// TIA Portal project "Milk Mixing 101" (V15.1)

(* hardware
DEVICE "S7-1200 station_1"  S7-1200 Station
   slot 0: "Rack_0"  S7-1200 Rack  Rack  V1.0
   slot 1: "PLC_1"  CPU 1214C AC/DC/Rly  6ES7 214-1BG40-0XB0  V4.2
DEVICE "PC-System_1"  SIMATIC PC station
   slot 0: "SIMATIC PC station"  Rail  SIMATIC PC-Station  V1.0
      slot 125: "Stationmanager"  Station_Manager  V6.0.4
   slot 1: "HMI_RT_1"  WinCC RT Advanced  6AV2 104-0xxxx-xxxx  15.1.0.0
      slot 33792: "Host interface"  Host interface
   slot 2: "IE general_1"  IE General  IE_CP  V8.2.0
*)

// ===== PLC "PLC_1"  CPU 1214C AC/DC/Rly =====

VAR_GLOBAL   // PLC tag table "Default tag table"
   "Auto_Start" AT %M0.0 : Bool;
   "Param_set" AT %M0.1 : Bool;
   "Timer_T123_ET" AT %MD0 : Time;
   "Filling_T123_Done" AT %M4.0 : Bool;
   "Filling_W1_Done" AT %M4.1 : Bool;
   "Mixing_Done" AT %M4.2 : Bool;
   "Pumping_Done" AT %M4.3 : Bool;
   "Pastorizing_Done" AT %M4.4 : Bool;
   "Filler_Done" AT %M4.5 : Bool;
   "MoveFork" AT %MD4 : DWord;
END_VAR

DATA_BLOCK "Recipe_Params"   // DB1
{ S7_Optimized_Access := 'TRUE' }
VERSION : 0.1
   VAR
      Flavour_Vol : Real;
      Milk_Vol : Real;
      Mixing_time : Time;
      Pastorizing_time : Time;
      Pastorizing_temp : Real;
      Filling_speed : Real;
      Flavour : Int;
   END_VAR
BEGIN
END_DATA_BLOCK

DATA_BLOCK "Devices"   // DB2
{ S7_Optimized_Access := 'TRUE' }
VERSION : 0.1
   VAR
      V11 : Bool;
      V12 : Bool;
      V13 : Bool;
      T1 : Bool;
      T2 : Bool;
      T3 : Bool;
      V21 : Bool;
      V22 : Bool;
      V23 : Bool;
      Mixer : Bool;
      W1 : Bool;
      V3 : Bool;
      Pump : Bool;
      V4 : Bool;
      Pastrorizer : Bool;
      v5 : Bool;
      Filler : Bool;
      Fork_Lift : Bool;
   END_VAR
BEGIN
END_DATA_BLOCK

DATA_BLOCK "SCADA_inputs"   // DB3
{ S7_Optimized_Access := 'TRUE' }
VERSION : 0.1
   VAR
      Start : Bool;
      Stop : Bool;
      Auto_On : Bool;
   END_VAR
BEGIN
END_DATA_BLOCK

DATA_BLOCK "Timer_ET"   // DB5
{ S7_Optimized_Access := 'TRUE' }
VERSION : 0.1
   VAR
      FillingTanks_ET : Time;
      FillingW1_ET : Time;
      MixingTimer_ET : Time;
      PumpingTimer_ET : Time;
      pastorizingTimer_ET : Time;
      FillerTimer_ET : Time;
   END_VAR
BEGIN
END_DATA_BLOCK

// folder: System blocks/Program resources

DATA_BLOCK "Filling_T1_2_3"   // DB4
{ S7_Optimized_Access := 'TRUE' }
AUTHOR : Simatic
FAMILY : IEC
NAME : IEC_TMR
VERSION : 1.0
// stored: InstanceOfName IEC_TIMER
"IEC_TIMER"
BEGIN
END_DATA_BLOCK

DATA_BLOCK "Filling_W1"   // DB6
{ S7_Optimized_Access := 'TRUE' }
AUTHOR : Simatic
FAMILY : IEC
NAME : IEC_TMR
VERSION : 1.0
// stored: InstanceOfName IEC_TIMER
"IEC_TIMER"
BEGIN
END_DATA_BLOCK

DATA_BLOCK "Mixing_timer"   // DB7
{ S7_Optimized_Access := 'TRUE' }
AUTHOR : Simatic
FAMILY : IEC
NAME : IEC_TMR
VERSION : 1.0
// stored: InstanceOfName IEC_TIMER
"IEC_TIMER"
BEGIN
END_DATA_BLOCK

DATA_BLOCK "Pumping_Timer"   // DB8
{ S7_Optimized_Access := 'TRUE' }
AUTHOR : Simatic
FAMILY : IEC
NAME : IEC_TMR
VERSION : 1.0
// stored: InstanceOfName IEC_TIMER
"IEC_TIMER"
BEGIN
END_DATA_BLOCK

DATA_BLOCK "Pastorizing_timer"   // DB9
{ S7_Optimized_Access := 'TRUE' }
AUTHOR : Simatic
FAMILY : IEC
NAME : IEC_TMR
VERSION : 1.0
// stored: InstanceOfName IEC_TIMER
"IEC_TIMER"
BEGIN
END_DATA_BLOCK

DATA_BLOCK "Filler_Timer"   // DB10
{ S7_Optimized_Access := 'TRUE' }
AUTHOR : Simatic
FAMILY : IEC
NAME : IEC_TMR
VERSION : 1.0
// stored: InstanceOfName IEC_TIMER
"IEC_TIMER"
BEGIN
END_DATA_BLOCK

DATA_BLOCK "Move_Fork"   // DB11
{ S7_Optimized_Access := 'TRUE' }
AUTHOR : Simatic
FAMILY : IEC
NAME : IEC_TMR
VERSION : 1.0
// stored: InstanceOfName IEC_TIMER
"IEC_TIMER"
BEGIN
END_DATA_BLOCK

// folder: (top level)

ORGANIZATION_BLOCK "Main"   // OB1, LAD, ProgramCycle
TITLE = "Main Program Sweep (Cycle)"
{ S7_Optimized_Access := 'TRUE' }
VERSION : 0.1
   VAR_INPUT
      Initial_Call : Bool;   // Initial call of this OB
      Remanence : Bool;   // =True, if remanent data are available
   END_VAR
BEGIN

REGION Network 1: Starting in Auto Mode
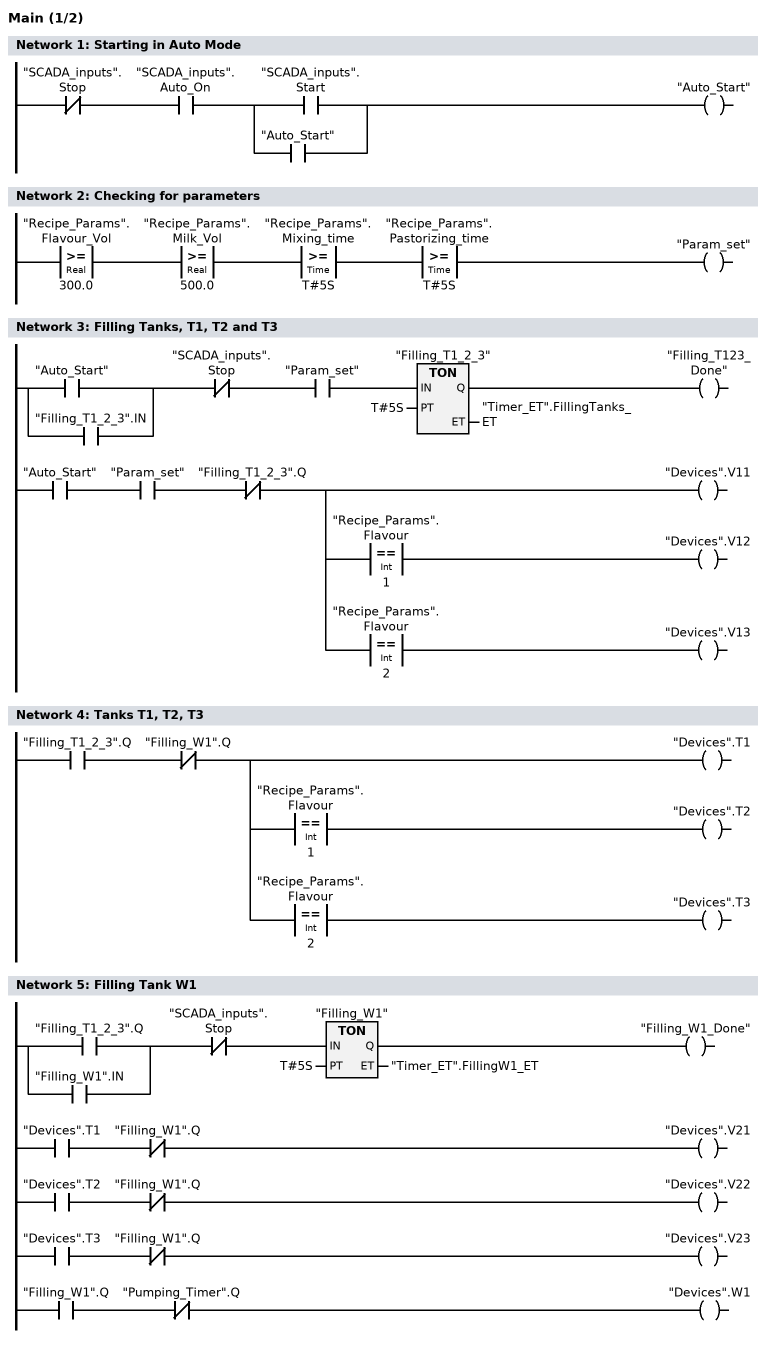
   RUNG wire#powerrail
      I_Contact( "SCADA_inputs".Stop )
      Contact( "SCADA_inputs".Auto_On )
      wire#w1
      Contact( "SCADA_inputs".Start )
      wire#w2
      Coil( "Auto_Start" )
   END_RUNG
   RUNG wire#w1
      Contact( "Auto_Start" )
   END_RUNG wire#w2
   // the same network as SCL:
   "Auto_Start" := NOT "SCADA_inputs".Stop AND "SCADA_inputs".Auto_On AND ("SCADA_inputs".Start OR "Auto_Start");
END_REGION

REGION Network 2: Checking for parameters
   RUNG wire#powerrail
      { S7_Templates := "SrcType := Real" } GE_Contact(in1 := "Recipe_Params".Flavour_Vol, in2 := 300.0)
      { S7_Templates := "SrcType := Real" } GE_Contact(in1 := "Recipe_Params".Milk_Vol, in2 := 500.0)
      { S7_Templates := "SrcType := Time" } GE_Contact(in1 := "Recipe_Params".Mixing_time, in2 := T#5S)
      { S7_Templates := "SrcType := Time" } GE_Contact(in1 := "Recipe_Params".Pastorizing_time, in2 := T#5S)
      Coil( "Param_set" )
   END_RUNG
   // the same network as SCL:
   "Param_set" := ("Recipe_Params".Flavour_Vol >= 300.0) AND ("Recipe_Params".Milk_Vol >= 500.0) AND ("Recipe_Params".Mixing_time >= T#5S) AND ("Recipe_Params".Pastorizing_time >= T#5S);
END_REGION

REGION Network 3: Filling Tanks, T1, T2 and T3
   "Filling_T1_2_3".TON(IN := ("Auto_Start" OR "Filling_T1_2_3".IN) AND NOT "SCADA_inputs".Stop AND "Param_set",
                        PT := T#5S,
                        ET => "Timer_ET".FillingTanks_ET);
   "Filling_T123_Done" := "Filling_T1_2_3".Q;
   "Devices".V11 := "Auto_Start" AND "Param_set" AND NOT "Filling_T1_2_3".Q;
   "Devices".V12 := "Devices".V11 AND ("Recipe_Params".Flavour = 1);
   "Devices".V13 := "Devices".V11 AND ("Recipe_Params".Flavour = 2);
END_REGION

REGION Network 4: Tanks T1, T2, T3
   RUNG wire#powerrail
      Contact( "Filling_T1_2_3".Q )
      I_Contact( "Filling_W1".Q )
      wire#w1
      Coil( "Devices".T1 )
   END_RUNG
   RUNG wire#w1
      { S7_Templates := "SrcType := Int" } EQ_Contact(in1 := "Recipe_Params".Flavour, in2 := 1)
      Coil( "Devices".T2 )
   END_RUNG
   RUNG wire#w1
      { S7_Templates := "SrcType := Int" } EQ_Contact(in1 := "Recipe_Params".Flavour, in2 := 2)
      Coil( "Devices".T3 )
   END_RUNG
   // the same network as SCL:
   "Devices".T1 := "Filling_T1_2_3".Q AND NOT "Filling_W1".Q;
   "Devices".T2 := "Devices".T1 AND ("Recipe_Params".Flavour = 1);
   "Devices".T3 := "Devices".T1 AND ("Recipe_Params".Flavour = 2);
END_REGION

REGION Network 5: Filling Tank W1
   "Filling_W1".TON(IN := ("Filling_T1_2_3".Q OR "Filling_W1".IN) AND NOT "SCADA_inputs".Stop,
                    PT := T#5S,
                    ET => "Timer_ET".FillingW1_ET);
   "Filling_W1_Done" := "Filling_W1".Q;
   "Devices".V21 := "Devices".T1 AND NOT "Filling_W1".Q;
   "Devices".V22 := "Devices".T2 AND NOT "Filling_W1".Q;
   "Devices".V23 := "Devices".T3 AND NOT "Filling_W1".Q;
   "Devices".W1 := "Filling_W1".Q AND NOT "Pumping_Timer".Q;
END_REGION

REGION Network 6: Mixing
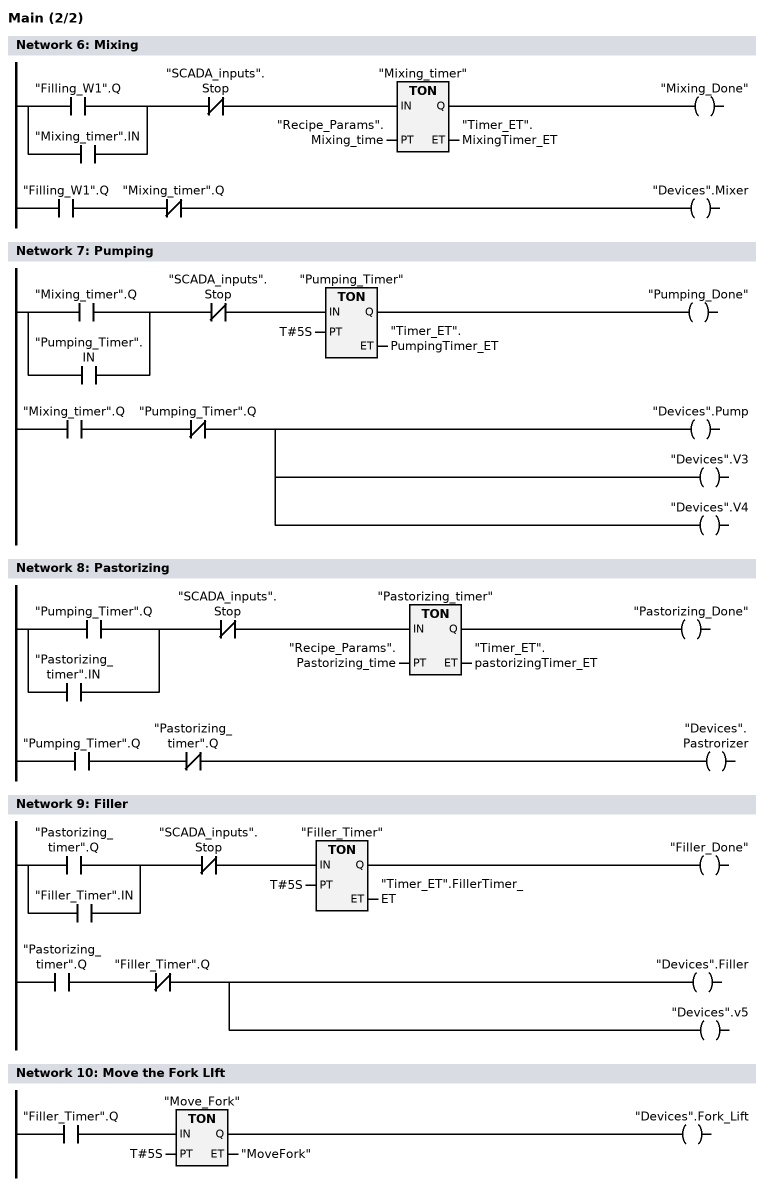
   "Mixing_timer".TON(IN := ("Filling_W1".Q OR "Mixing_timer".IN) AND NOT "SCADA_inputs".Stop,
                      PT := "Recipe_Params".Mixing_time,
                      ET => "Timer_ET".MixingTimer_ET);
   "Mixing_Done" := "Mixing_timer".Q;
   "Devices".Mixer := "Filling_W1".Q AND NOT "Mixing_timer".Q;
END_REGION

REGION Network 7: Pumping
   "Pumping_Timer".TON(IN := ("Mixing_timer".Q OR "Pumping_Timer".IN) AND NOT "SCADA_inputs".Stop,
                       PT := T#5S,
                       ET => "Timer_ET".PumpingTimer_ET);
   "Pumping_Done" := "Pumping_Timer".Q;
   "Devices".Pump := "Mixing_timer".Q AND NOT "Pumping_Timer".Q;
   "Devices".V3 := "Devices".Pump;
   "Devices".V4 := "Devices".Pump;
END_REGION

REGION Network 8: Pastorizing
   "Pastorizing_timer".TON(IN := ("Pumping_Timer".Q OR "Pastorizing_timer".IN) AND NOT "SCADA_inputs".Stop,
                           PT := "Recipe_Params".Pastorizing_time,
                           ET => "Timer_ET".pastorizingTimer_ET);
   "Pastorizing_Done" := "Pastorizing_timer".Q;
   "Devices".Pastrorizer := "Pumping_Timer".Q AND NOT "Pastorizing_timer".Q;
END_REGION

REGION Network 9: Filler
   "Filler_Timer".TON(IN := ("Pastorizing_timer".Q OR "Filler_Timer".IN) AND NOT "SCADA_inputs".Stop,
                      PT := T#5S,
                      ET => "Timer_ET".FillerTimer_ET);
   "Filler_Done" := "Filler_Timer".Q;
   "Devices".Filler := "Pastorizing_timer".Q AND NOT "Filler_Timer".Q;
   "Devices".v5 := "Devices".Filler;
END_REGION

REGION Network 10: Move the Fork LIft
   "Move_Fork".TON(IN := "Filler_Timer".Q, PT := T#5S, ET => "MoveFork");
   "Devices".Fork_Lift := "Move_Fork".Q;
END_REGION
END_ORGANIZATION_BLOCK

(* ===== HMI "HMI_RT_1" =====
system functions are stored by id; their names below are inferred from use
connection "HMI_Connection_1": ETHERNET, S7_1200_OMS

HMI tags "Default tag table"
   "Recipe_Params_Flavour" : Int = PLC Recipe_Params.Flavour, 1 s
   "Recipe_Params_Flavour_Vol" : Real = PLC Recipe_Params.Flavour_Vol, 1 s
   "Recipe_Params_Milk_Vol" : Real = PLC Recipe_Params.Milk_Vol, 1 s
   "Recipe_Params_Mixing_time" : Time = PLC Recipe_Params.Mixing_time, 1 s
   "Recipe_Params_Pastorizing_time" : Time = PLC Recipe_Params.Pastorizing_time, 1 s
   "Recipe_Params_Pastorizing_temp" : Real = PLC Recipe_Params.Pastorizing_temp, 1 s
   "Recipe_Params_Filling_speed" : Real = PLC Recipe_Params.Filling_speed, 1 s
   "SCADA_inputs_Start" : Bool = PLC SCADA_inputs.Start, 1 s
   "SCADA_inputs_Stop" : Bool = PLC SCADA_inputs.Stop, 1 s
   "SCADA_inputs_Auto_On" : Bool = PLC SCADA_inputs.Auto_On, 1 s
   "Devices_V11" : Bool = PLC Devices.V11, 1 s
   "Devices_V12" : Bool = PLC Devices.V12, 1 s
   "Devices_V13" : Bool = PLC Devices.V13, 1 s
   "Devices_T1" : Bool = PLC Devices.T1, 1 s
   "Devices_T2" : Bool = PLC Devices.T2, 1 s
   "Devices_T3" : Bool = PLC Devices.T3, 1 s
   "Devices_V21" : Bool = PLC Devices.V21, 1 s
   "Devices_V22" : Bool = PLC Devices.V22, 1 s
   "Devices_V23" : Bool = PLC Devices.V23, 1 s
   "Devices_Mixer" : Bool = PLC Devices.Mixer, 1 s
   "Devices_W1" : Bool = PLC Devices.W1, 1 s
   "Devices_V3" : Bool = PLC Devices.V3, 1 s
   "Devices_Pump" : Bool = PLC Devices.Pump, 1 s
   "Devices_V4" : Bool = PLC Devices.V4, 1 s
   "Devices_Pastrorizer" : Bool = PLC Devices.Pastrorizer, 1 s
   "Devices_v5" : Bool = PLC Devices.v5, 1 s
   "Devices_Filler" : Bool = PLC Devices.Filler, 1 s
   "MoveFork" : DWord = PLC MoveFork AT %MD4, 1 s
   "Timer_ET_FillingW1_ET" : Time = PLC Timer_ET.FillingW1_ET, 1 s
   "Auto_Start" : Bool = PLC Auto_Start AT %M0.0, 1 s

text list "Flavour": 1 'Strawberry'; 2 'Chocolate'

screen "Main_Screen" 1920x1068
   TextField "Text field_1" at 647,26 size 456x34; Text 'MILK MIXING SYSTEM'
   SymbolLibrary "Symbol library_1" at 52,135 size 108x126
   SymbolLibrary "Symbol library_2" at 254,136 size 108x126
   SymbolLibrary "Symbol library_3" at 459,136 size 108x126
   SymbolLibrary "Symbol library_4" at 66,359 size 85x71
      Appearance <- "Devices_T1"
   SymbolLibrary "Symbol library_5" at 267,356 size 85x71
      Appearance <- "Devices_T2"
   SymbolLibrary "Symbol library_6" at 471,360 size 85x71
      Appearance <- "Devices_T3"
   SymbolLibrary "Symbol library_7" at 98,262 size 16x99
      Appearance <- "Devices_V11"
   SymbolLibrary "Symbol library_8" at 300,262 size 16x99
      Appearance <- "Devices_V12"
   SymbolLibrary "Symbol library_9" at 507,261 size 16x99
      Appearance <- "Devices_V13"
   SymbolLibrary "Symbol library_10" at 77,292 size 38x41
      Appearance <- "Devices_V11"
   SymbolLibrary "Symbol library_11" at 280,290 size 38x41
      Appearance <- "Devices_V12"
   SymbolLibrary "Symbol library_12" at 487,292 size 38x41
      Appearance <- "Devices_V13"
   SymbolLibrary "Symbol library_13" at 211,552 size 201x153
      Appearance <- "Devices_W1"
   SymbolLibrary "Symbol library_14" at 100,425 size 16x84
      Appearance <- "Devices_V21"
   SymbolLibrary "Symbol library_15" at 302,426 size 16x130
      Appearance <- "Devices_V22"
   SymbolLibrary "Symbol library_16" at 506,430 size 16x76
      Appearance <- "Devices_V23"
   SymbolLibrary "Symbol library_17" at 384,517 size 103x16
      Appearance <- "Devices_V23"
   SymbolLibrary "Symbol library_18" at 133,518 size 83x16
      Appearance <- "Devices_V21"
   SymbolLibrary "Symbol library_19" at 352,516 size 33x35
   SymbolLibrary "Symbol library_20" at 213,517 size 29x38
   SymbolLibrary "Symbol library_21" at 99,505 size 35x27
   SymbolLibrary "Symbol library_22" at 486,502 size 36x30
   SymbolLibrary "Symbol library_23" at 525,809 size 101x89
      Appearance <- "Devices_Pump"
   SymbolLibrary "Symbol library_25" at 299,704 size 23x120
      Appearance <- "Devices_V3"
   SymbolLibrary "Symbol library_26" at 339,842 size 188x17
      Appearance <- "Devices_V3"
   SymbolLibrary "Symbol library_24" at 416,812 size 43x49
      Appearance <- "Devices_V3"
   SymbolLibrary "Symbol library_27" at 299,823 size 42x37
   SymbolLibrary "Symbol library_28" at 822,414 size 120x120
      Appearance <- "Devices_Pastrorizer"
   SymbolLibrary "Symbol library_29" at 713,502 size 18x301
      Appearance <- "Devices_V4"
   SymbolLibrary "Symbol library_30" at 626,818 size 59x20
   SymbolLibrary "Symbol library_31" at 751,466 size 76x19
      Appearance <- "Devices_V4"
   SymbolLibrary "Symbol library_32" at 712,466 size 39x39
   SymbolLibrary "Symbol library_33" at 685,801 size 49x36
   SymbolLibrary "Symbol library_34" at 762,436 size 43x49
      Appearance <- "Devices_V4"
   SymbolLibrary "Symbol library_35" at 858,678 size 120x120
      Appearance <- "Devices_Filler"
   SymbolLibrary "Symbol library_36" at 869,522 size 21x157
      Appearance <- "Devices_v5"
   SymbolLibrary "Symbol library_37" at 832,582 size 64x35
      Appearance <- "Devices_v5"
   SymbolLibrary "Symbol library_38" at 973,755 size 239x43
   SymbolLibrary "Symbol library_39" at 1206,691 size 120x120
      HorizontalMovement <- "MoveFork"
   Switch "Switch_1" at 1130,109 size 108x55; CaptionText 'MODE'; TextOff 'MANUAL'; TextOn 'AUTO'
      on SwitchOn: SetBit("SCADA_inputs_Auto_On")
      on SwitchOff: ResetBit("SCADA_inputs_Auto_On")
   Button "Button_1" at 1285,129 size 96x32; TextOff 'START'
      on Press: SetBit("SCADA_inputs_Start")
      on Release: ResetBit("SCADA_inputs_Start")
   Button "Button_2" at 1437,130 size 96x32; TextOff 'STOP'
      on Press: SetBit("SCADA_inputs_Stop")
      on Release: ResetBit("SCADA_inputs_Stop")
   TextField "Text field_2" at 1221,197 size 321x27; Text 'Recipe Parameter'
   TextField "Text field_3" at 1149,278 size 115x22; Text 'Flavour'
   TextField "Text field_4" at 1137,338 size 179x22; Text 'Flavour Volume'
   TextField "Text field_5" at 1140,386 size 159x22; Text 'Milk Volume'
   TextField "Text field_6" at 1138,426 size 155x22; Text 'Mixing Time'
   TextField "Text field_7" at 1134,470 size 185x22; Text 'Pastorizing Time'
   TextField "Text field_8" at 1135,515 size 198x22; Text 'Pastorizing Temp'
   TextField "Text field_9" at 1141,560 size 182x22; Text 'Filling Speed'
   SymbolicIOField "Symbolic I/O field_1" at 1294,277 size 142x33; TextOff '0'; TextOn '1'; TextList "Flavour"
      ProcessValue <- "Recipe_Params_Flavour"
      Visibility <- "Auto_Start"
   IOField "I/O field_1" at 1296,333 size 96x32; FormatPattern 9999
      ProcessValue <- "Recipe_Params_Flavour_Vol"
      Visibility <- "Auto_Start"
   IOField "I/O field_2" at 1296,382 size 96x32; FormatPattern 9999
      ProcessValue <- "Recipe_Params_Milk_Vol"
      Visibility <- "Auto_Start"
   IOField "I/O field_3" at 1296,422 size 96x32; FormatPattern 99999
      ProcessValue <- "Recipe_Params_Mixing_time"
      Visibility <- "Auto_Start"
   IOField "I/O field_4" at 1297,466 size 96x32; FormatPattern 99999
      ProcessValue <- "Recipe_Params_Pastorizing_time"
      Visibility <- "Auto_Start"
   IOField "I/O field_5" at 1298,511 size 96x32; FormatPattern 9999
      ProcessValue <- "Recipe_Params_Pastorizing_temp"
      Visibility <- "Auto_Start"
   IOField "I/O field_6" at 1297,558 size 96x32; FormatPattern 9999
      ProcessValue <- "Recipe_Params_Filling_speed"
      Visibility <- "Auto_Start"
   TextField "Text field_10" at 1415,337 size 53x22; Text 'ltr'
   TextField "Text field_11" at 1412,382 size 56x22; Text 'ltr'
   TextField "Text field_12" at 1410,426 size 77x22; Text 'ms'
   TextField "Text field_13" at 1408,476 size 87x22; Text 'ms'
   TextField "Text field_14" at 1413,516 size 81x22; Text 'c'
   TextField "Text field_15" at 1399,560 size 177x22; Text 'Bottle/min'
   TextField "Text field_16" at 43,300 size 35x22; Text 'V11'
   TextField "Text field_17" at 245,300 size 35x22; Text 'V12'
   TextField "Text field_18" at 453,302 size 35x22; Text 'V13'
   TextField "Text field_19" at 100,376 size 24x22; Text 'T1'
   TextField "Text field_20" at 302,372 size 24x22; Text 'T2'
   TextField "Text field_21" at 498,376 size 24x22; Text 'T3'
   SymbolLibrary "Symbol library_40" at 73,454 size 47x35
      Appearance <- "Devices_V21"
   SymbolLibrary "Symbol library_41" at 272,457 size 47x35
      Appearance <- "Devices_V22"
   SymbolLibrary "Symbol library_42" at 478,457 size 47x35
      Appearance <- "Devices_V23"
   TextField "Text field_22" at 40,461 size 35x22; Text 'V21'
   TextField "Text field_23" at 237,464 size 35x22; Text 'V22'
   TextField "Text field_24" at 443,467 size 35x22; Text 'V23'
   TextField "Text field_25" at 289,657 size 30x22; Text 'W1'
   SymbolLibrary "Symbol library_43" at 240,519 size 73x75
      Appearance <- "Devices_Mixer"
   TextField "Text field_26" at 257,600 size 48x22; Text 'Mixer'
   TextField "Text field_27" at 423,790 size 25x22; Text 'V3'
   TextField "Text field_28" at 770,415 size 25x22; Text 'V4'
   TextField "Text field_29" at 546,787 size 46x22; Text 'Pump'
   TextField "Text field_30" at 827,393 size 195x22; Text 'Pastorizer'
   TextField "Text field_31" at 807,590 size 25x22; Text 'V5'
   TextField "Text field_32" at 912,694 size 133x22; Text 'Filler'
   TextField "Text field_33" at 1153,716 size 132x22; Text 'Fork Lift'
   Bar "Bar_1" at 410,550 size 63x164; MinimumValue 0; MaximumValue 5000
      ProcessValue <- "Timer_ET_FillingW1_ET"
   TextField "Text field_34" at 61,100 size 125x22; Text 'MILK'
   TextField "Text field_35" at 261,104 size 170x22; Text 'STRAWBERRY'
   TextField "Text field_36" at 485,106 size 185x22; Text 'CHOCOLATE'
   TextField "Text field_37" at 1508,279 size 154x22; Text 'Text'
   TextField "Text field_38" at 1507,343 size 139x22; Text 'Text'
   TextField "Text field_39" at 1507,383 size 157x22; Text 'Text'
   TextField "Text field_40" at 1503,431 size 151x22; Text 'Text'
   TextField "Text field_41" at 1506,486 size 142x22; Text 'Text'
*)